         IF #statExternalStopDetected = FALSE THEN
           // handle usual internal stop reaction
           IF #instMC_GROUPSTOP.Busy = FALSE THEN
             // check TO Kinematics to have stopped successfully
             IF (#to_Kinematics.StatusWord.%X12 = TRUE)                        // TO Kinematics with constant velocity
               AND (#to_Kinematics.StatusPath.Velocity = 0.0)                  // TO Kinematics path velocity 0.0
               AND (#to_Kinematics.StatusMotionQueue.NumberOfCommands = 0)     // MotionQueue deleted completely
               AND (#instMC_GROUPSTOP.Done = TRUE)
             THEN
               #statStateMachine := #STOPPED_STATE;
             ELSE
               // set execute trigger for MC_GroupStop
               #statExecGroupStop := TRUE;
             END_IF;
           ELSE
             // Added FR: 08.04.2019
             // stop conditions fulfilled without GroupStop executed successfully (done <> TRUE, busy = TRUE)
             IF (#to_Kinematics.StatusWord.%X12 = TRUE)                        // TO Kinematics with constant velocity
               AND (#to_Kinematics.StatusWord.%X6 = TRUE)                      // no jobs active on TO Kinematics
               AND (#to_Kinematics.StatusWord.%X16 = FALSE)                    // TO Kinematics not stopping anymore ==> GroupStop done
               AND (#to_Kinematics.StatusPath.Velocity = 0.0)                  // TO Kinematics path velocity 0.0
               AND (#to_Kinematics.StatusMotionQueue.NumberOfCommands = 0)     // MotionQueue deleted completely
             THEN
               #statStateMachine := #STOPPED_STATE;
             END_IF;
           END_IF;

         ELSE
           // handle external stop
           IF (#to_Kinematics.StatusWord.%X12 = TRUE)                        // TO Kinematics with constant velocity
             AND (#to_Kinematics.StatusWord.%X6 = TRUE)                      // no jobs active on TO Kinematics
             AND (#to_Kinematics.StatusWord.%X16 = FALSE)                    // TO Kinematics not stopping anymore ==> GroupStop done
             AND (#to_Kinematics.StatusPath.Velocity = 0.0)                  // TO Kinematics path velocity 0.0
             AND (#to_Kinematics.StatusMotionQueue.NumberOfCommands = 0)     // MotionQueue deleted completely
           THEN
             #statStateMachine := #STOPPED_STATE;
             // reset bit for detection of external stop triggered
             #statExternalStopDetected := FALSE;
           END_IF;
         END_IF;

       END_IF;

     END_REGION STOPPING


     // state reached when GroupStop is executed ==> do nothing when stopped
     REGION STOPPED_STATE
       IF #statStateMachine = #STOPPED_STATE
         // AND #statDebugState = TRUE
       THEN
         // reset  variable for single step debugging of states
         #statDebugState := FALSE;

         #statExecGroupStop := FALSE;

         // check for MC_GroupStop to be finished or inactive
         IF #instMC_GROUPSTOP.Busy = FALSE THEN
           #statStatus := #STATUS_COMMAND_ABORTED;
         END_IF;

         // Check stopMode if desync from conveyor shall be executed
         IF (#tempStopMode = 10 OR #tempStopMode = 11) AND #statActualTrackedOCS <> 0 THEN
           #statStateMachine := #DESYNC_CONVEYOR;
           #statStatus := #STATUS_DESYNC_CONVEYOR;
         END_IF;

       END_IF;
     END_REGION STOPPED_STATE


     REGION STOP_DESYNC_CONVEYOR
       IF #statStateMachine = #DESYNC_CONVEYOR
         // AND #statDebugState = TRUE
       THEN
         // Check if linear cmd is done or not busy anymore
         IF #instMC_MoveLinAbs[#statFBCounterLin].Done
           OR (#instMC_MoveLinAbs[#statFBCounterLin].Busy = FALSE
           AND #statExecLinCmds[#statFBCounterLin] = TRUE)
         THEN
           #statExecLinCmds[#statFBCounterLin] := FALSE;
           #statStatus := #STATUS_COMMAND_ABORTED;
         END_IF;

         // Check if stop is not active at kinematics --> Linear cmd is not rejected
         IF #to_Kinematics.StatusWord.%X16 = FALSE AND #statStatus <> #STATUS_COMMAND_ABORTED THEN
           // Execute linear cmd in wcs
           #statAbsolutePosition[1] := #to_Kinematics.TcpInWcs.x.Position;
           #statAbsolutePosition[2] := #to_Kinematics.TcpInWcs.y.Position;
           #statAbsolutePosition[3] := #to_Kinematics.TcpInWcs.z.Position;
           #statAbsolutePosition[4] := #to_Kinematics.TcpInWcs.a.Position;
           #statExecLinCmds[#statFBCounterLin] := true;
           #pathDataElementPreBuf.cmdCoordinates.coordSystem := "CS_WCS";
           #pathDataElementPreBuf.cmdParameters.pathDynamics.velocity := -1;
           #pathDataElementPreBuf.cmdParameters.pathDynamics.acceleration := -1;
           #pathDataElementPreBuf.cmdParameters.pathDynamics.deceleration := -1;
           #pathDataElementPreBuf.cmdParameters.pathDynamics.jerk := -1;
           #pathDataElementPreBuf.cmdParameters.dynamicAdaption := 0; // DA must be off
           #pathDataElementPreBuf.cmdParameters.bufferMode := 1;
         END_IF;

       END_IF;
     END_REGION STOP_DESYNC_CONVEYOR


     // wait for requesting new command when MotionQueue is busy with executed commands
     REGION QUEUE_BUSY
       IF #statStateMachine = #QUEUE_BUSY THEN // check for new command already waiting to be executed
         // check for MotionQueue to be ready buffering new commands from PathDataPreBuffered
         IF #to_Kinematics.StatusMotionQueue.NumberOfCommands < #to_Kinematics.MotionQueue.MaxNumberOfCommands
           AND #instMC_GROUPSTOP.Busy = FALSE
         THEN
           // MotionQueue ready ==> continue execution
           // receive new command when buffer is ready for new command
           #statStateMachine := #RECEIVE_CMD;
         ELSE
           // set status information, do nothing, wait for buffer to be ready again
           #statStatus := #STATUS_PATHMOTION_BUFFER_BUSY;
         END_IF;
       END_IF;
     END_REGION QUEUE_BUSY


     // state reached when error occured ==> do nothing when error occured
     REGION ERROR_STATE
       IF #statStateMachine = #ERROR_STATE
         // AND #statDebugState = TRUE
       THEN
         // reset  variable for single step debugging of states
         #statDebugState := FALSE;

         // reset all execute triggers for motion commands in case of error
         FOR #tempCtr := 1 TO #LKINCTRL_MAX_NUMBER_OF_CMDS_LIN DO
           #statExecLinCmds[#tempCtr] := FALSE;
           #statExecCircCmds[#tempCtr] := FALSE;
           #statExecMoveDirectCmds[#tempCtr] := FALSE;
         END_FOR;

         FOR #tempCtr := 1 TO #LKINCTRL_MAX_NUMBER_OF_CMDS_TRACKCONV DO
           #statExecTrackConv[#tempCtr] := FALSE;
         END_FOR;
       END_IF;
     END_REGION ERROR_STATE

   END_REGION STATE_MACHINE

   REGION CHECK_FINISHED_CMDs
     //----------------------------------------------------------------------------------------------
     // FB Execution & Analysis
     //----------------------------------------------------------------------------------------------
     // Only check finished cmds if FB is still busy & commands shall be executed
     IF #statBusy
       AND (#statStateMachine < #INTERRUPTING // all states below 70
       OR #statStateMachine = #CONTINUEING // or state = 77
       OR #statStateMachine = #CONTINUED) // or state = 78
     THEN
       // Init temporary variables
       #tempCmdDone := FALSE;
       #tempActiveInstance := 0;
       #tempCmdType := #statStoreExecuteBuffer.bufferElement[#statStoreExecuteBuffer.activeBufferElement].MotionFBNo;

       // Check motionFBNo
       IF #tempCmdType <= -1 THEN
         #tempActiveInstance := 0;
       ELSIF #tempCmdType = "LKINCTRL_CMD_WAIT_TIME" THEN
         #tempActiveInstance := 0;
       ELSIF #tempCmdType = "LKINCTRL_CMD_FLAG_ONLY" THEN
         #tempActiveInstance := 0;
       ELSIF #tempCmdType > "LKINCTRL_CMD_WAIT_TIME" AND #tempCmdType <= "LKINCTRL_CMD_WAIT_TIME" + #LKINCTRL_MAX_NUMBER_OF_CMDS_TRACKCONV THEN
         // TrackConveyor command (101..103)
         #tempActiveInstance := #tempCmdType - "LKINCTRL_CMD_WAIT_TIME";
         #tempCmdType := "LKINCTRL_MC_TRACKCONVEYORBELT";
       ELSE
         // MotionFBNo is actual MC command
         // --> Calculate type and active instance
         IF #tempCmdType MOD #LKINCTRL_EXECUTEBUFFER_LENGTH <> 0 THEN
           #tempCmdType := (#tempCmdType / #LKINCTRL_EXECUTEBUFFER_LENGTH);
         ELSE
           #tempCmdType := (#tempCmdType / #LKINCTRL_EXECUTEBUFFER_LENGTH) - 1;
         END_IF;
         // Calc active MC instance 
         #tempActiveInstance := #statStoreExecuteBuffer.bufferElement[#statStoreExecuteBuffer.activeBufferElement].MotionFBNo - #LKINCTRL_EXECUTEBUFFER_LENGTH * #tempCmdType;
         // Increase type once more to fit lower case
         #tempCmdType += 1;
       END_IF;

       // Reset debug variables
       #statDebugMessage := '';
       #statDebugFaultyValue := 0;

       CASE #tempCmdType OF
         "LKINCTRL_CMD_FLAG_ONLY": // FlagOnly
           // check for flagOnly command to have been 'executed' (activeCmdNo has been written to output for at least one cycle)
           // eventually replace by this
           IF #statStoreExecuteBuffer.bufferElement[#statStoreExecuteBuffer.activeBufferElement].setNumber = #writtenActiveCmdNo THEN
             // reset bit for flagOnly command is 'active'
             #statExecuteFlagOnlyCmd := FALSE;
             #tempCmdDone := TRUE;
           END_IF;

         1:  // Linear
           // check active MotionFB to be done
           IF #instMC_MoveLinAbs[#tempActiveInstance].#Done THEN
             // reset execute trigger at MotionFB.execute if MotionFB is done
             #statExecLinCmds[#tempActiveInstance] := FALSE;
             // Set temp to signal cmd is done
             #tempCmdDone := TRUE;
           END_IF;

         2:  // Circular
           IF #instMC_MoveCircAbs[#tempActiveInstance].Done THEN
             // reset execute trigger at MotionFB.execute if MotionFB is done
             #statExecCircCmds[#tempActiveInstance] := FALSE;
             // Set temp to signal cmd is done
             #tempCmdDone := TRUE;
           END_IF;

         3: // MoveDirect
           IF #instMC_MoveDirectAbs[#tempActiveInstance].Done THEN
             // reset execute trigger at MotionFB.execute if MotionFB is done
             #statExecMoveDirectCmds[#tempActiveInstance] := FALSE;
             // Set temp to signal cmd is done
             #tempCmdDone := TRUE;
           END_IF;

         "LKINCTRL_MC_TRACKCONVEYORBELT":
           IF #instMC_TrackConveyor[#tempActiveInstance].Done
             OR (#to_Kinematics.StatusConveyor[#instMC_TrackConveyor[#tempActiveInstance].CoordSystem].TrackingState = 1) // Done is sometimes not set, so check TrackingState also
           THEN
             // reset execute trigger at MotionFB.execute if MotionFB is done
             #statExecTrackConv[#tempActiveInstance] := FALSE;
             // Set temp to signal cmd is done
             #tempCmdDone := TRUE;
           END_IF;

         "LKINCTRL_CMD_WAIT_TIME": // WaitTime
           IF #instIEC_Timer_waitTime.Q = TRUE THEN
             // reset trigger for WAIT_TIME when timer is done
             #statExecWaitTime := FALSE;
             #tempCmdDone := TRUE;
             // Set remainingDistance to 0.0 if done --> sometimes 1 would still appear because of dataType conversion error
             #remainingDistanceActCmd := 0.0;
           END_IF;

         ELSE  // Undefined cmd
           #statDebugMessage := 'motionFBNo (Done) out of range 1...20';
           #statDebugFaultyValue := #statStoreExecuteBuffer.bufferElement[#statStoreExecuteBuffer.activeBufferElement].MotionFBNo;
       END_CASE;

       // Check if the active cmd is done
       IF #tempCmdDone THEN
         // Reset blending radius calculation
         #statBlendingRadius := -1;

         // Check if cmd was last command to be executed
         IF #statStoreExecuteBuffer.activeBufferElement = #statStoreExecuteBuffer.lastBufferElement THEN
           // Set status to pathmotion finished
           #statStatus := #STATUS_PATHMOTION_FINISHED;
         ELSE
           // Increase activeBufferElement when not finished
           // check statStoreExecureBuffer counter for active elements not to exceed statStoreExecuteBuffer.bufferElements[1..LKINCTRL_EXECUTEBUFFER_LENGTH] length
           IF #statStoreExecuteBuffer.activeBufferElement < #LKINCTRL_EXECUTEBUFFER_LENGTH THEN
             // increase statStoreExecureBuffer counter for active elements
             #statStoreExecuteBuffer.activeBufferElement := #statStoreExecuteBuffer.activeBufferElement + 1;
           ELSE
             // reset statStoreExecureBuffer counter for active elements
             #statStoreExecuteBuffer.activeBufferElement := 1;
           END_IF;

           // check for new activeBufferElement to be flagOnly command
           IF #statStoreExecuteBuffer.bufferElement[#statStoreExecuteBuffer.activeBufferElement].MotionFBNo = "LKINCTRL_CMD_FLAG_ONLY" THEN
             // set 'active' bit for flagOnly command
             #statExecuteFlagOnlyCmd := TRUE;
           ELSE
             #statExecuteFlagOnlyCmd := FALSE;
           END_IF;

           // increment activeCmdLogger pointer
           IF #statDebugExecCmdLogger.activeCmdLoggerElement < #CONST_LENGTH_DATALOGGER THEN
             #statDebugExecCmdLogger.activeCmdLoggerElement := #statDebugExecCmdLogger.activeCmdLoggerElement + 1;
           ELSE
             #statDebugExecCmdLogger.activeCmdLoggerElement := 1;
           END_IF;
         END_IF;
       END_IF;
     END_IF;
   END_REGION CHECK_FINISHED_CMDs

   REGION CALL_MC_CMDs

     REGION LIN_CIRC_MOVEDIRECT_CMDs
       // FB Execution cyclically to update FB outputs
       FOR #tempFBInstCtr := 1 TO #LKINCTRL_MAX_NUMBER_OF_CMDS_LIN DO
         // execute all linear  motion command FBs with set control variables in every cycle
         #instMC_MoveLinAbs[#tempFBInstCtr](AxesGroup := #to_Kinematics,
                                            Execute := #statExecLinCmds[#tempFBInstCtr],
                                            Position := #statAbsolutePosition,
                                            Velocity := #pathDataElementPreBuf.cmdParameters.pathDynamics.velocity,
                                            Acceleration := #pathDataElementPreBuf.cmdParameters.pathDynamics.acceleration,
                                            Deceleration := #pathDataElementPreBuf.cmdParameters.pathDynamics.deceleration,
                                            Jerk := #pathDataElementPreBuf.cmdParameters.pathDynamics.jerk,
                                            DirectionA := #pathDataElementPreBuf.cmdParameters.orientationDirection,
                                            CoordSystem := #pathDataElementPreBuf.cmdCoordinates.coordSystem,
                                            BufferMode := #pathDataElementPreBuf.cmdParameters.bufferMode,
                                            TransitionParameter := #pathDataElementPreBuf.cmdParameters.transitionParameters,
                                            DynamicAdaption := #pathDataElementPreBuf.cmdParameters.dynamicAdaption);
         // check all FBs for occurred error in every cycle 
         IF #instMC_MoveLinAbs[#tempFBInstCtr].Error
           AND (#statStatus.%X15 = FALSE) // Check if other error was already set
           AND #statStatus <> #STATUS_PATHMOTION_STOPPING // Check if instance is aborted because of stop
         THEN
           // exclude error from MC_GroupStop ==> handled in stop routine
           IF #instMC_MoveLinAbs[#tempFBInstCtr].ErrorId <> 16#80CD THEN
             #statStatus := #ERR_LINEAR_CMD;
           END_IF;
           #statSubfunctionStatus := #instMC_MoveLinAbs[#tempFBInstCtr].ErrorId;
           #diagnostics.#faultFBNumber := #tempFBInstCtr;
           #diagnostics.#faultSetNumber := #statStoreExecuteBuffer.bufferElement[#statStoreExecuteBuffer.activeBufferElement].setNumber;
           #diagnostics.#faultPathDataName := #statStoreExecuteBuffer.bufferElement[#statStoreExecuteBuffer.activeBufferElement].pathDataName;
         END_IF;
       END_FOR;

       FOR #tempFBInstCtr := 1 TO #LKINCTRL_MAX_NUMBER_OF_CMDS_CIRC DO
         // execute all circular  motion command FBs with set control variables in every cycle
         #instMC_MoveCircAbs[#tempFBInstCtr](AxesGroup := #to_Kinematics,
                                             Execute := #statExecCircCmds[#tempFBInstCtr],
                                             CircMode := #pathDataElementPreBuf.cmdParameters.circleParameters.circMode,
                                             AuxPoint := #statAuxPoint,
                                             EndPoint := #statEndPoint,
                                             PathChoice := #pathDataElementPreBuf.cmdParameters.circleParameters.pathChoice,
                                             CirclePlane := #pathDataElementPreBuf.cmdParameters.circleParameters.circlePlane,
                                             Radius := #pathDataElementPreBuf.cmdParameters.circleParameters.radius,
                                             Arc := #pathDataElementPreBuf.cmdParameters.circleParameters.arc,
                                             Velocity := #pathDataElementPreBuf.cmdParameters.pathDynamics.velocity,
                                             Acceleration := #pathDataElementPreBuf.cmdParameters.pathDynamics.acceleration,
                                             Deceleration := #pathDataElementPreBuf.cmdParameters.pathDynamics.deceleration,
                                             Jerk := #pathDataElementPreBuf.cmdParameters.pathDynamics.jerk,
                                             DirectionA := #pathDataElementPreBuf.cmdParameters.orientationDirection,
                                             CoordSystem := #pathDataElementPreBuf.cmdCoordinates.coordSystem,
                                             BufferMode := #pathDataElementPreBuf.cmdParameters.bufferMode,
                                             TransitionParameter := #pathDataElementPreBuf.cmdParameters.transitionParameters,
                                             DynamicAdaption := #pathDataElementPreBuf.cmdParameters.dynamicAdaption);
         // check all FBs for occurred error in every cycle 
         IF #instMC_MoveCircAbs[#tempFBInstCtr].Error
           AND (#statStatus.%X15 = FALSE) // Check if other error was already set
           AND #statStatus <> #STATUS_PATHMOTION_STOPPING // Check if instance is aborted because of stop
         THEN
           // exclude error from MC_GroupStop
           IF #instMC_MoveCircAbs[#tempFBInstCtr].ErrorId <> 16#80CD THEN
             #statStatus := #ERR_CIRCULAR_CMD;
           END_IF;
           #statSubfunctionStatus := #instMC_MoveCircAbs[#tempFBInstCtr].ErrorId;
           #diagnostics.faultFBNumber := #tempFBInstCtr + #LKINCTRL_EXECUTEBUFFER_LENGTH;
           #diagnostics.#faultSetNumber := #statStoreExecuteBuffer.bufferElement[#statStoreExecuteBuffer.activeBufferElement].setNumber;
           #diagnostics.#faultPathDataName := #statStoreExecuteBuffer.bufferElement[#statStoreExecuteBuffer.activeBufferElement].pathDataName;
         END_IF;
       END_FOR;

       FOR #tempFBInstCtr := 1 TO #LKINCTRL_MAX_NUMBER_OF_CMDS_MOVEDIRECT DO
         // execute all move direct motion command FBs with set control variables in every cycle
         #instMC_MoveDirectAbs[#tempFBInstCtr](AxesGroup := #to_Kinematics,
                                               Execute := #statExecMoveDirectCmds[#tempFBInstCtr],
                                               Position := #statAbsolutePosition,
                                               VelocityFactor := #pathDataElementPreBuf.cmdParameters.pathDynamics.velocity,
                                               AccelerationFactor := #pathDataElementPreBuf.cmdParameters.pathDynamics.acceleration,
                                               DecelerationFactor := #pathDataElementPreBuf.cmdParameters.pathDynamics.deceleration,
                                               JerkFactor := #pathDataElementPreBuf.cmdParameters.pathDynamics.jerk,
                                               LinkConstellation := #pathDataElementPreBuf.cmdParameters.moveDirectParameters.linkConstellation,
                                               PositionMode := #pathDataElementPreBuf.cmdParameters.moveDirectParameters.positionMode,
                                               DirectionA := #pathDataElementPreBuf.cmdParameters.orientationDirection,
                                               CoordSystem := #pathDataElementPreBuf.cmdCoordinates.coordSystem,
                                               BufferMode := #pathDataElementPreBuf.cmdParameters.bufferMode,
                                               TransitionParameter := #pathDataElementPreBuf.cmdParameters.transitionParameters);
         // check all FBs for occurred error in every cycle 
         IF #instMC_MoveDirectAbs[#tempFBInstCtr].Error
           AND (#statStatus.%X15 = FALSE) // Check if other error was already set
           AND #statStatus <> #STATUS_PATHMOTION_STOPPING // Check if instance is aborted because of stop
         THEN
           // exclude error from MC_GroupStop ==> handled in stop routine
           IF #instMC_MoveDirectAbs[#tempFBInstCtr].ErrorId <> 16#80CD THEN
             #statStatus := #ERR_MOVEDIRECT_CMD;
           END_IF;
           #statSubfunctionStatus := #instMC_MoveDirectAbs[#tempFBInstCtr].ErrorId;
           #diagnostics.#faultFBNumber := #tempFBInstCtr + 2 * #LKINCTRL_EXECUTEBUFFER_LENGTH;
           #diagnostics.#faultSetNumber := #statStoreExecuteBuffer.bufferElement[#statStoreExecuteBuffer.activeBufferElement].setNumber;
           #diagnostics.#faultPathDataName := #statStoreExecuteBuffer.bufferElement[#statStoreExecuteBuffer.activeBufferElement].pathDataName;
         END_IF;
       END_FOR;
     END_REGION LIN_CIRC_MOVEDIRECT_CMDs


     REGION TRACK_CONVEYOR
       FOR #tempFBInstCtr := 1 TO #LKINCTRL_MAX_NUMBER_OF_CMDS_TRACKCONV DO
         // execute all track conveyor motion command FBs with set control variables in every cycle
         #instMC_TrackConveyor[#tempFBInstCtr].Execute := #statExecTrackConv[#tempFBInstCtr];

         IF TypeOfDB(#statConveyorBeltAxis[#tempFBInstCtr]) = TO_POSITIONINGAXIS THEN
           "LKinCtrl_CallMC_TrackConv_PosAxis"(posAxis := #statConveyorBeltAxis[#tempFBInstCtr],
                                               axesGroup := #to_Kinematics,
                                               instTrackConveyorBelt := #instMC_TrackConveyor[#tempFBInstCtr]);

         ELSIF TypeOfDB(#statConveyorBeltAxis[#tempFBInstCtr]) = TO_SYNCHRONOUSAXIS THEN
           "LKinCtrl_CallMC_TrackConv_SyncAxis"(syncAxis := #statConveyorBeltAxis[#tempFBInstCtr],
                                                axesGroup := #to_Kinematics,
                                                instTrackConveyorBelt := #instMC_TrackConveyor[#tempFBInstCtr]);

         ELSIF TypeOfDB(#statConveyorBeltAxis[#tempFBInstCtr]) = TO_EXTERNALENCODER THEN
           "LKinCtrl_CallMC_TrackConv_ExtEncoder"(extEncoder := #statConveyorBeltAxis[#tempFBInstCtr],
                                                  axesGroup := #to_Kinematics,
                                                  instTrackConveyorBelt := #instMC_TrackConveyor[#tempFBInstCtr]);

         ELSIF TypeOfDB(#statConveyorBeltAxis[#tempFBInstCtr]) = TO_LeadingAxisProxy THEN
           "LKinCtrl_CallMC_TrackConv_LeadingAxisProxy"(leadingAxisProxy := #statConveyorBeltAxis[#tempFBInstCtr],
                                                        axesGroup := #to_Kinematics,
                                                        instTrackConveyorBelt := #instMC_TrackConveyor[#tempFBInstCtr]);

         ELSE
           ; // Error wrong axis type or no axis connected ?!
         END_IF;

         // check all FBs for occurred error in every cycle 
         IF #instMC_TrackConveyor[#tempFBInstCtr].Error
           AND (#statStatus.%X15 = FALSE) // Check if other error was already set
           AND #statStatus <> #STATUS_PATHMOTION_STOPPING // Check if instance is aborted because of stop
         THEN
           // exclude error from MC_GroupStop ==> handled in stop routine
           IF #instMC_TrackConveyor[#tempFBInstCtr].ErrorId <> 16#80CD THEN
             #statStatus := #ERR_TRACKCONVEYOR_CMD;
           END_IF;
           #statSubfunctionStatus := #instMC_TrackConveyor[#tempFBInstCtr].ErrorId;
           #diagnostics.#faultFBNumber := #tempFBInstCtr + "LKINCTRL_CMD_WAIT_TIME";
           #diagnostics.#faultSetNumber := #statStoreExecuteBuffer.bufferElement[#statStoreExecuteBuffer.activeBufferElement].setNumber;
           #diagnostics.#faultPathDataName := #statStoreExecuteBuffer.bufferElement[#statStoreExecuteBuffer.activeBufferElement].pathDataName;
         END_IF;
       END_FOR;

     END_REGION TRACK_CONVEYOR


     REGION MC_CTRL_CMDs

       #instMC_GROUPINTERRUPT(AxesGroup := #to_Kinematics,
                              Execute := #statExecGroupInterrupt,
                              Mode := 0);
       // error detection and signaling
       IF #instMC_GROUPINTERRUPT.Error THEN
         #statSubfunctionStatus := #instMC_GROUPCONTINUE.ErrorId;
         // set status for error evaluation ==> statError will be set in output section
         #statStatus := #ERR_GROUPINTERRUPT_FAILED;
       END_IF;

       // Reset execute of interrupt
       IF #instMC_GROUPINTERRUPT.Done OR #instMC_GROUPINTERRUPT.CommandAborted THEN
         #instMC_GROUPINTERRUPT(AxesGroup := #to_Kinematics,
                                Execute := FALSE);
       END_IF;

       #instMC_GROUPCONTINUE(AxesGroup := #to_Kinematics,
                             Execute := #statExecGroupContinue);
       // error detection and signaling
       IF #instMC_GROUPCONTINUE.Error THEN
         #statSubfunctionStatus := #instMC_GROUPCONTINUE.ErrorId;
         // set status for error evaluation ==> statError will be set in output section
         #statStatus := #ERR_GROUPCONTINUE_FAILED;
       END_IF;

       // Reset execute of continue
       IF #instMC_GROUPCONTINUE.Done THEN
         #instMC_GROUPCONTINUE(AxesGroup := #to_Kinematics,
                               Execute := FALSE);
       END_IF;

       // Check for correct stop mode
       CASE #tempStopMode OF
         0, 1: // normal stopMode
           #tempStopMode := #tempStopMode;
         10: // stopMode with stop of conveyor (path dynamics)
           #tempStopMode := 0;
         11: // stopMode with stop of conveyor (maximum dynamics)
           #tempStopMode := 1;
         ELSE
           // Invalid stop mode specification 
           // Use maximum dynamics
           #tempStopMode := 1;
       END_CASE;

       #instMC_GROUPSTOP(AxesGroup := #to_Kinematics,
                         Execute := #statExecGroupStop,
                         Mode := #tempStopMode);
       // error detection and signaling
       IF #instMC_GROUPSTOP.Error THEN
         #statSubfunctionStatus := #instMC_GROUPSTOP.ErrorId;
         // set status for error evaluation ==> statError will be set in output section
         #statStatus := #ERR_GROUPSTOP_FAILED;
       END_IF;

       // call WAIT_TIME
       #instIEC_Timer_waitTime(IN := #statExecWaitTime,
                               PT := #statWaitTime);

     END_REGION MC_CTRL_CMDs

   END_REGION CALL_MC_CMDs

   REGION CHECK_TO_KINEMATICS_STATE

     // check TO_Kinematics for pending errors
     IF #to_Kinematics.StatusWord.%X1 = TRUE THEN
       // only copy statusWords to outputs in case of error
       #diagnostics.kinematicsStatusWord := #to_Kinematics.StatusWord;
       #diagnostics.kinematicsErrorWord := #to_Kinematics.ErrorWord;

       // set status
       #statStatus := #ERR_TO_KINEMATIC_ERROR;
     END_IF;

     IF #to_Kinematics.StatusWord.%X16 = TRUE
       AND #statStateMachine <> #STOPPING
       AND #statStateMachine <> #STOPPED_STATE
       AND #statStateMachine <> #DESYNC_CONVEYOR
       AND #statStateMachine <> #ERROR_STATE
       AND #tempStop = FALSE
     THEN
       // set bit for detection of external stop
       #statExternalStopDetected := TRUE;
       // set state machine
       #statStateMachine := #STOPPING;
       #statStatus := #STATUS_PATHMOTION_EXT_STOPPING;
     END_IF;

     // Check if conveyor is tracked
     FOR #tempCtr := 1 TO 3 DO
       #statActualTrackedOCS := 0;
       IF #to_Kinematics.StatusConveyor[#tempCtr].TrackingState = 3 THEN
         #statActualTrackedOCS := DINT_TO_SINT(#tempCtr);
         EXIT;
       END_IF;
     END_FOR;

   END_REGION CHECK_TO_KINEMATICS_STATE

   REGION OUTPUTS
     //----------------------------------------------------------------------------------------------
     // Write ouputs and error handling
     //----------------------------------------------------------------------------------------------
     REGION ACTIVE_CMD
       // Only check active cmds if FB is still busy
       IF #statBusy THEN
         // check to_kinematics to reset active
         IF #to_Kinematics.StatusWord.%X8 = FALSE
           AND #to_Kinematics.StatusWord.%X9 = FALSE
           AND #to_Kinematics.StatusWord.%X11 = FALSE
         THEN
           // reset active output
           #statActive := FALSE;
         END_IF;

         // Init temporary variables
         #tempActiveInstance := 0;
         #tempCmdType := #statStoreExecuteBuffer.bufferElement[#statStoreExecuteBuffer.activeBufferElement].MotionFBNo;

         // Check motionFBNo
         IF #tempCmdType <= -1 THEN
           #tempActiveInstance := 0;
         ELSIF #tempCmdType = "LKINCTRL_CMD_WAIT_TIME" THEN
           #tempActiveInstance := 0;
         ELSIF #tempCmdType = "LKINCTRL_CMD_FLAG_ONLY" THEN
           #tempActiveInstance := 0;
         ELSIF #tempCmdType > "LKINCTRL_CMD_WAIT_TIME" AND #tempCmdType <= "LKINCTRL_CMD_WAIT_TIME" + #LKINCTRL_MAX_NUMBER_OF_CMDS_TRACKCONV THEN
           // TrackConveyor command (101..103)
           #tempActiveInstance := #tempCmdType - "LKINCTRL_CMD_WAIT_TIME";
           #tempCmdType := "LKINCTRL_MC_TRACKCONVEYORBELT";
         ELSE
           // MotionFBNo is actual MC command
           // --> Calculate type and active instance
           IF #tempCmdType MOD #LKINCTRL_EXECUTEBUFFER_LENGTH <> 0 THEN
             #tempCmdType := (#tempCmdType / #LKINCTRL_EXECUTEBUFFER_LENGTH);
           ELSE
             #tempCmdType := (#tempCmdType / #LKINCTRL_EXECUTEBUFFER_LENGTH) - 1;
           END_IF;
           // Calc active MC instance 
           #tempActiveInstance := #statStoreExecuteBuffer.bufferElement[#statStoreExecuteBuffer.activeBufferElement].MotionFBNo - #LKINCTRL_EXECUTEBUFFER_LENGTH * #tempCmdType;
           // Increase type once more to fit lower case
           #tempCmdType += 1;
         END_IF;

         // Reset debug variables
         #statDebugMessage := '';
         #statDebugFaultyValue := 0;

         CASE #tempCmdType OF
           "LKINCTRL_CMD_FLAG_ONLY": // FlagOnly
             ; // Do not change active state

           1:  // Linear
             // Always update remainingDistance
             #remainingDistanceActCmd := #instMC_MoveLinAbs[#tempActiveInstance].RemainingDistance;
             // check MotionFB to be active
             IF #instMC_MoveLinAbs[#tempActiveInstance].Active
               // 2019/09/17 - added JR: additional condition only for immediately done commands after flagOnly
               OR (#instMC_MoveLinAbs[#tempActiveInstance].Done
               // 2019/09/18 - added JR: neglect condition if next command is WAIT_TIME
               AND #statStateMachine <> #EXEC_WAIT_TIME)
             THEN
               // write activeCmd specific data to outputs
               #statActive := TRUE;
             END_IF;


           2:  // Circular
             // Always update remainingDistance
             #remainingDistanceActCmd := #instMC_MoveCircAbs[#tempActiveInstance].RemainingDistance;
             IF #instMC_MoveCircAbs[#tempActiveInstance].Active
               // 2019/09/18 - added JR: additional condition for immediately done commands after flagOnly
               OR (#instMC_MoveCircAbs[#tempActiveInstance].Done
               // 2019/09/18 - added JR: neglect condition if next command is WAIT_TIME
               AND #statStateMachine <> #EXEC_WAIT_TIME)
             THEN
               // write activeCmd specific data to outputs
               #statActive := TRUE;
             END_IF;

           3: // MoveDirect
             // -------------------------
             // Calculate own remDistance
             // TODO:
             // - When target is MCS then use Trafo FB to calc cartesian target
             // -------------------------
             // Get coord system
             #tempCtr := DINT_TO_INT(#statDebugExecCmdLogger.loggerElement[#statDebugExecCmdLogger.activeCmdLoggerElement].executedCmd.coordSystem);

             IF #SPTP_REMAINING_DIST AND #tempCtr <> "CS_MCS" THEN
               // Deactivate blending calculation if setting is off
               IF #SPTP_APPROX_BLENDING = FALSE THEN
                 #statBlendingRadius := 0;
               END_IF;

               // Only do this if blending is not calculated already for this command 
               IF #statBlendingRadius = -1 THEN
                 // Calculate blending radius
                 // Get blending setting and target of following command
                 IF #statDebugExecCmdLogger.activeCmdLoggerElement <> #CONST_LENGTH_DATALOGGER THEN
                   IF #statDebugExecCmdLogger.activeCmdLoggerElement + 1 <> #statDebugExecCmdLogger.writeCmdLoggerElement THEN
                     #tempBlending[1] := #statDebugExecCmdLogger.loggerElement[#statDebugExecCmdLogger.activeCmdLoggerElement + 1].executedCmd.bufferMode;
                     #tempBlending[2] := #statDebugExecCmdLogger.loggerElement[#statDebugExecCmdLogger.activeCmdLoggerElement + 1].executedCmd.transitionParameter;
                     #tempCalc[1] := #statDebugExecCmdLogger.loggerElement[#statDebugExecCmdLogger.activeCmdLoggerElement + 1].executedCmd.coordinateX;
                     #tempCalc[2] := #statDebugExecCmdLogger.loggerElement[#statDebugExecCmdLogger.activeCmdLoggerElement + 1].executedCmd.coordinateY;
                     #tempCalc[3] := #statDebugExecCmdLogger.loggerElement[#statDebugExecCmdLogger.activeCmdLoggerElement + 1].executedCmd.coordinateZ;
                     "LKinCtrl_FrameTrans"(coordSystem := #tempCtr,
                                           coordSystemOld := #statDebugExecCmdLogger.loggerElement[#statDebugExecCmdLogger.activeCmdLoggerElement + 1].executedCmd.coordSystem,
                                           OCSFrames := #statOCSFrames,
                                           position := #tempCalc);
                   END_IF;
                 ELSE
                   IF 1 <> #statDebugExecCmdLogger.writeCmdLoggerElement THEN
                     #tempBlending[1] := #statDebugExecCmdLogger.loggerElement[1].executedCmd.bufferMode;
                     #tempBlending[2] := #statDebugExecCmdLogger.loggerElement[1].executedCmd.transitionParameter;
                     #tempCalc[1] := #statDebugExecCmdLogger.loggerElement[1].executedCmd.coordinateX;
                     #tempCalc[2] := #statDebugExecCmdLogger.loggerElement[1].executedCmd.coordinateY;
                     #tempCalc[3] := #statDebugExecCmdLogger.loggerElement[1].executedCmd.coordinateZ;
                     "LKinCtrl_FrameTrans"(coordSystem := #tempCtr,
                                           coordSystemOld := #statDebugExecCmdLogger.loggerElement[1].executedCmd.coordSystem,
                                           OCSFrames := #statOCSFrames,
                                           position := #tempCalc);
                   END_IF;
                 END_IF;

                 // Check blending settings
                 IF (#tempBlending[1] = "BM_BLENDING_LOW" OR #tempBlending[1] = "BM_BLENDING_HIGH") AND #tempBlending[2] <> 0.0 THEN
                   // Calc blending from the two targets
                   // Calc length of second command
                   #tempCalc[1] -= #statDebugExecCmdLogger.loggerElement[#statDebugExecCmdLogger.activeCmdLoggerElement].executedCmd.coordinateX;
                   #tempCalc[2] -= #statDebugExecCmdLogger.loggerElement[#statDebugExecCmdLogger.activeCmdLoggerElement].executedCmd.coordinateY;
                   #tempCalc[3] -= #statDebugExecCmdLogger.loggerElement[#statDebugExecCmdLogger.activeCmdLoggerElement].executedCmd.coordinateZ;
                   // Calculate length of vector (actual to next)
                   #tempBlending[3] := SQRT(#tempCalc[1] * #tempCalc[1] + #tempCalc[2] * #tempCalc[2] + #tempCalc[3] * #tempCalc[3]);
                 ELSE
                   #statBlendingRadius := 0;
                 END_IF;

                 // TODO: Get last target for blending radius calculation
                 IF #statDebugExecCmdLogger.activeCmdLoggerElement <> 1 THEN
                   IF #statDebugExecCmdLogger.activeCmdLoggerElement - 1 <> #statDebugExecCmdLogger.writeCmdLoggerElement THEN
                     #tempCalc[1] := #statDebugExecCmdLogger.loggerElement[#statDebugExecCmdLogger.activeCmdLoggerElement - 1].executedCmd.coordinateX;
                     #tempCalc[2] := #statDebugExecCmdLogger.loggerElement[#statDebugExecCmdLogger.activeCmdLoggerElement - 1].executedCmd.coordinateY;
                     #tempCalc[3] := #statDebugExecCmdLogger.loggerElement[#statDebugExecCmdLogger.activeCmdLoggerElement - 1].executedCmd.coordinateZ;
                     "LKinCtrl_FrameTrans"(coordSystem := #tempCtr,
                                           coordSystemOld := #statDebugExecCmdLogger.loggerElement[#statDebugExecCmdLogger.activeCmdLoggerElement - 1].executedCmd.coordSystem,
                                           OCSFrames := #statOCSFrames,
                                           position := #tempCalc);
                   END_IF;
                 ELSE
                   IF #CONST_LENGTH_DATALOGGER <> #statDebugExecCmdLogger.writeCmdLoggerElement THEN
                     #tempCalc[1] := #statDebugExecCmdLogger.loggerElement[#CONST_LENGTH_DATALOGGER].executedCmd.coordinateX;
                     #tempCalc[2] := #statDebugExecCmdLogger.loggerElement[#CONST_LENGTH_DATALOGGER].executedCmd.coordinateY;
                     #tempCalc[3] := #statDebugExecCmdLogger.loggerElement[#CONST_LENGTH_DATALOGGER].executedCmd.coordinateZ;
                     "LKinCtrl_FrameTrans"(coordSystem := #tempCtr,
                                           coordSystemOld := #statDebugExecCmdLogger.loggerElement[1].executedCmd.coordSystem,
                                           OCSFrames := #statOCSFrames,
                                           position := #tempCalc);
                   END_IF;
                 END_IF;

                 // Calc length of first command 
                 #tempCalc[1] := #statDebugExecCmdLogger.loggerElement[#statDebugExecCmdLogger.activeCmdLoggerElement].executedCmd.coordinateX - #tempCalc[1];
                 #tempCalc[2] := #statDebugExecCmdLogger.loggerElement[#statDebugExecCmdLogger.activeCmdLoggerElement].executedCmd.coordinateY - #tempCalc[2];
                 #tempCalc[3] := #statDebugExecCmdLogger.loggerElement[#statDebugExecCmdLogger.activeCmdLoggerElement].executedCmd.coordinateZ - #tempCalc[3];
                 // Calculate length of vector (last to actual)
                 #tempBlending[4] := SQRT(#tempCalc[1] * #tempCalc[1] + #tempCalc[2] * #tempCalc[2] + #tempCalc[3] * #tempCalc[3]);
               END_IF;

               // Assign target value
               #tempCalc[1] := #statDebugExecCmdLogger.loggerElement[#statDebugExecCmdLogger.activeCmdLoggerElement].executedCmd.coordinateX;
               #tempCalc[2] := #statDebugExecCmdLogger.loggerElement[#statDebugExecCmdLogger.activeCmdLoggerElement].executedCmd.coordinateY;
               #tempCalc[3] := #statDebugExecCmdLogger.loggerElement[#statDebugExecCmdLogger.activeCmdLoggerElement].executedCmd.coordinateZ;
               // Substract kinematics position
               IF #tempCtr = "CS_WCS" THEN
                 #tempCalc[1] -= #to_Kinematics.TcpInWcs.x.Position;
                 #tempCalc[2] -= #to_Kinematics.TcpInWcs.y.Position;
                 #tempCalc[3] -= #to_Kinematics.TcpInWcs.z.Position;
               ELSE
                 #tempCalc[1] -= #to_Kinematics.TcpInOcs[#tempCtr].x.Position;
                 #tempCalc[2] -= #to_Kinematics.TcpInOcs[#tempCtr].y.Position;
                 #tempCalc[3] -= #to_Kinematics.TcpInOcs[#tempCtr].z.Position;
               END_IF;

               // Calculate length of vector
               #remainingDistanceActCmd := SQRT(#tempCalc[1] * #tempCalc[1] + #tempCalc[2] * #tempCalc[2] + #tempCalc[3] * #tempCalc[3]);

               // Check which command is shorter distance
               IF #statBlendingRadius = -1 THEN
                 IF #tempBlending[2] < 0.0 THEN // Transition parameter 
                   // Check which command is shorter     //Last target to current       //Current target to next
                   #statBlendingRadius := MIN_LREAL(IN1 := #tempBlending[4] / 2.0, IN2 := #tempBlending[3] / 2.0);
                 ELSE
                   // Check which setting is the shortest
                   #statBlendingRadius := MIN_LREAL(IN1 := #tempBlending[4] / 2.0, IN2 := #tempBlending[3] / 2.0, IN3 := #tempBlending[2]);
                 END_IF;
               END_IF;

               // Calculate remaining distance
               #remainingDistanceActCmd -= #statBlendingRadius;
               IF #remainingDistanceActCmd < 0.0 THEN // Avoid negative values
                 #remainingDistanceActCmd := 0.0;
               END_IF;

             ELSE
               // Always update remainingDistance
               #remainingDistanceActCmd := #instMC_MoveDirectAbs[#tempActiveInstance].ExecutionTimeStatus;
             END_IF;

             // Check active state
             IF #instMC_MoveDirectAbs[#tempActiveInstance].Active
               // 2019/09/18 - added JR: additional condition for immediately done commands after flagOnly
               OR (#instMC_MoveDirectAbs[#tempActiveInstance].Done
               // 2019/09/18 - added JR: neglect condition if next command is WAIT_TIME
               AND #statStateMachine <> #EXEC_WAIT_TIME)
             THEN
               // write activeCmd specific data to outputs
               #statActive := TRUE;
             END_IF;

           "LKINCTRL_MC_TRACKCONVEYORBELT": // TrackConveoyrBelt
             IF #instMC_TrackConveyor[#tempActiveInstance].Busy // No active output at instance --> Use busy
               // 2019/09/18 - added JR: additional condition for immediately done commands after flagOnly
               OR (#instMC_TrackConveyor[#tempActiveInstance].Done
               // 2019/09/18 - added JR: neglect condition if next command is WAIT_TIME
               AND #statStateMachine <> #EXEC_WAIT_TIME)
             THEN
               #statActive := TRUE;
             END_IF;

           "LKINCTRL_CMD_WAIT_TIME": // WaitTime
             // Reset active output
             #statActive := FALSE;
             // Calculate remainingDistance
             IF #instIEC_Timer_waitTime.ET <> t#0ms THEN
               #remainingDistanceActCmd := TIME_TO_UDINT(#statWaitTime - #instIEC_Timer_waitTime.ET);
             ELSIF #instIEC_Timer_waitTime.ET = t#0ms AND #instIEC_Timer_waitTime.IN = TRUE THEN
               #remainingDistanceActCmd := TIME_TO_UDINT(#statWaitTime);
             END_IF;

           ELSE  // Undefined cmd
             #statActive := FALSE;
             #remainingDistanceActCmd := 0.0;
             #statDebugMessage := 'motionFBNo (active) out of range 1...20';
             #statDebugFaultyValue := #statStoreExecuteBuffer.bufferElement[#statStoreExecuteBuffer.activeBufferElement].MotionFBNo;
         END_CASE;

         // Double check if to Kinematics is interrupted
         IF #to_Kinematics.StatusWord.%X17 = TRUE AND #instMC_GROUPCONTINUE.Busy = FALSE THEN
             #statActive := FALSE;
         END_IF;

         // write activeCmd specific data to outputs
         // Only update outputs if command is actually active to avoid issues with flagMode 5 & 10
         IF #statActive
           OR #tempCmdType = "LKINCTRL_CMD_WAIT_TIME"
           OR #tempCmdType = "LKINCTRL_CMD_FLAG_ONLY"
         THEN
           #activePathDataName := #statStoreExecuteBuffer.bufferElement[#statStoreExecuteBuffer.activeBufferElement].pathDataName;
           #activePathDataIdentifier := #statStoreExecuteBuffer.bufferElement[#statStoreExecuteBuffer.activeBufferElement].pathDataIdentifier;
           #statActiveCmdNo := #statStoreExecuteBuffer.bufferElement[#statStoreExecuteBuffer.activeBufferElement].setNumber;
         END_IF;
       END_IF;
     END_REGION ACTIVE_CMD


     REGION STATUS_EVALUATION
       // Write outputs
       IF (#statStatus.%X15 = TRUE) AND (#statError = FALSE) AND (#statBusy = TRUE) THEN // Error occurred (#statStatus is 16#8000 to 16#FFFF)
         #statDone := FALSE;
         #statBusy := FALSE;
         #statActive := FALSE;
         #statCommandAborted := FALSE;
         #statCmdExecuted := FALSE;
         #statError := TRUE;
         #statWaitTimeActive := FALSE;
         // Write diagnostics
         #diagnostics.stateMachine := #statStateMachine;
         #diagnostics.status := #statStatus;
         #diagnostics.motionFBstatus := #statSubfunctionStatus;
         #statStateMachine := #ERROR_STATE;

       ELSIF ((#statStatus = #STATUS_CMD_EXECUTED) AND (#statStatus <> #STATUS_WAIT_TIME_ACTIVE)) AND (#statDone = FALSE) THEN // command executed to MotionQueue, wait for next execution or end of path reached
         #statDone := FALSE;
         #statCommandAborted := FALSE;
         #statError := FALSE;
         #statCmdExecuted := TRUE;
         #statStateMachine := #NO_PROCESSING; // Switch state machine to "no processing"

       ELSIF (#statStatus = #STATUS_PATHMOTION_FINISHED) AND (#statDone = FALSE) THEN // Execution finished without errors
         #statDone := TRUE;
         #statBusy := FALSE;
         #statCommandAborted := FALSE;
         #statError := FALSE;
         #statWaitTimeActive := FALSE;
         #statStateMachine := #NO_PROCESSING; // Switch state machine to "no processing"
         #remainingDistanceActCmd := 0.0; // Reset remaining distance when done --> SPTP stays at 1.0, so a reset is necessary

       ELSIF (#statStatus = #STATUS_COMMAND_ABORTED) AND (#statCommandAborted = FALSE) THEN // Commanded functionality has been aborted by another command
         #statDone := FALSE;
         #statBusy := FALSE;
         #statCommandAborted := TRUE;
         #statError := FALSE;
         #statCmdExecuted := FALSE;
         #statWaitTimeActive := FALSE;
         // Write diagnostics
         #diagnostics.stateMachine := #statStateMachine;
         #diagnostics.status := #statStatus;
         #diagnostics.motionFBstatus := #statSubfunctionStatus;
         #statStateMachine := #NO_PROCESSING;

       ELSIF (#tempExecute = FALSE) AND (#tempStop = FALSE) AND ((#statDone = TRUE) OR (#statError = TRUE) OR (#statCommandAborted = TRUE)) THEN // Reset outputs
         #statDone := FALSE;
         #statBusy := FALSE;
         #statActive := FALSE;
         #statCommandAborted := FALSE;
         #statError := FALSE;
         #statCmdExecuted := FALSE;
         #statWaitTimeActive := FALSE;
         #statStatus := #STATUS_NO_CALL;
         // added FR: 2019/04/18 - set state machine to no processing, when ending FB
         #statStateMachine := #NO_PROCESSING;
       END_IF;

       // Write static values to outputs
       #done := #statDone;
       #busy := #statBusy;
       #active := #statActive;
       #activeCmdNo := #statActiveCmdNo;
       #waitTimeActive := #statWaitTimeActive;
       #commandAborted := #statCommandAborted;
       #error := #statError;
       #diagnostics.status := #statStatus;
       #cmdExecuted := #statCmdExecuted;
     END_REGION STATUS_EVALUATION

   END_REGION OUTPUTS
   // =================================================================================================================
   // End of Function Block: LKinCtrl_MC_ExecuteKinMotionCmd
   // =================================================================================================================
END_FUNCTION_BLOCK

// folder: LKinCtrl_Blocks/LKinCtrl_SubBlocks/LKinCtrl_ContOffsetBlocks

FUNCTION "LKinCtrl_OffsetContour" : "LKinCtrl_typeCOffReturn"   // FC35050, SCL
TITLE = LKinCtrl_OffsetContour
{ S7_Optimized_Access := 'TRUE' }
AUTHOR : tech.team.motioncontrol@siemens.com
FAMILY : LKinCtrl